// TIA Portal project "Pesteproject" (V15.1) (continued)
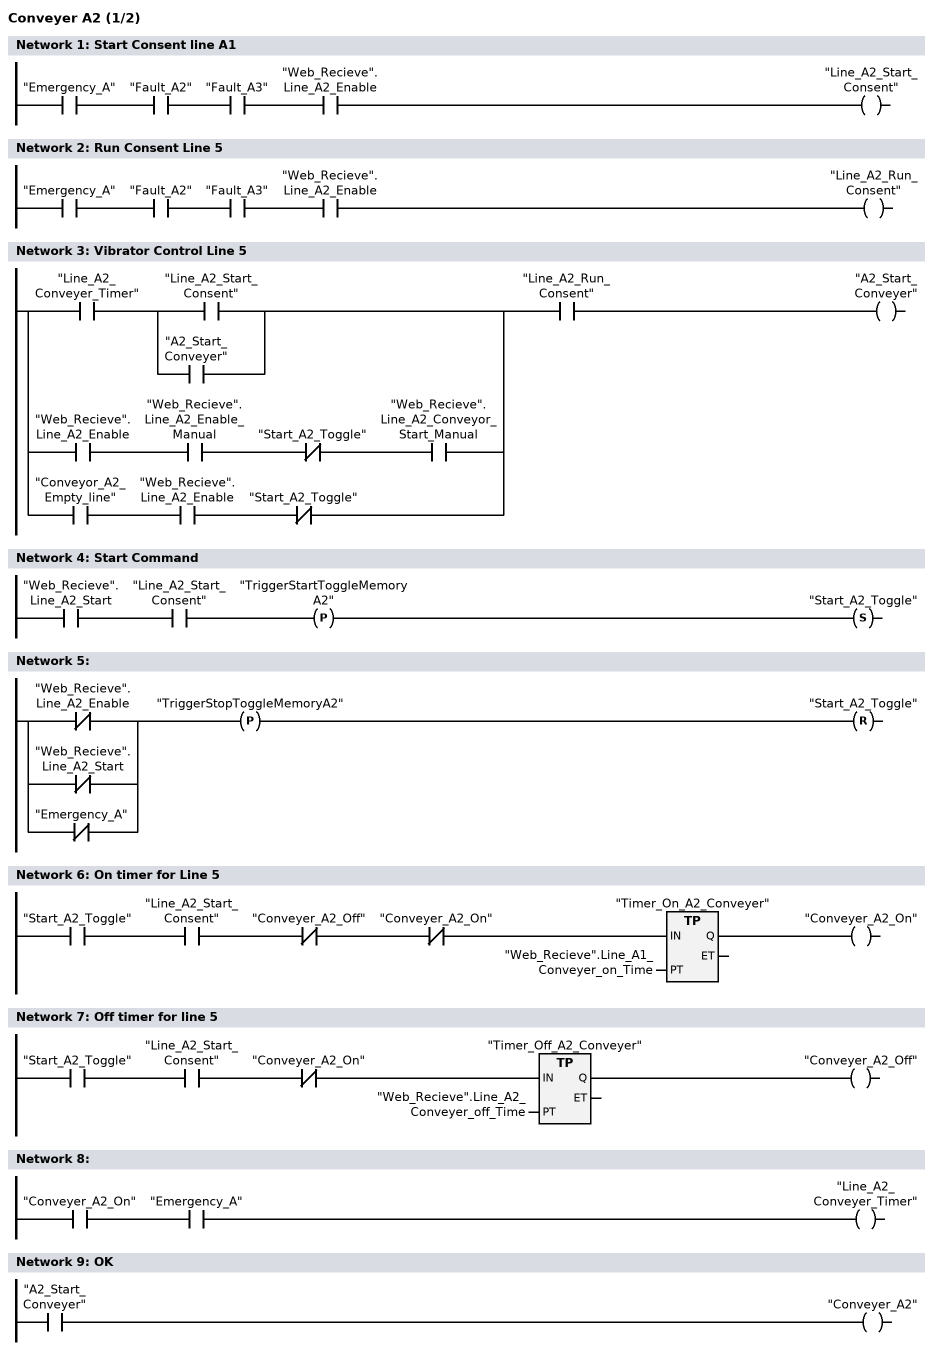
   RUNG wire#powerrail
      Contact( "Emergency_A" )
      Contact( "Fault_A2" )
      Contact( "Fault_A3" )
      Contact( "Web_Recieve".Line_A2_Enable )
      Coil( "Line_A2_Start_Consent" )
   END_RUNG
   // the same network as SCL:
   "Line_A2_Start_Consent" := "Emergency_A" AND "Fault_A2" AND "Fault_A3" AND "Web_Recieve".Line_A2_Enable;
END_REGION

REGION Network 2: Run Consent Line 5
   RUNG wire#powerrail
      Contact( "Emergency_A" )
      Contact( "Fault_A2" )
      Contact( "Fault_A3" )
      Contact( "Web_Recieve".Line_A2_Enable )
      Coil( "Line_A2_Run_Consent" )
   END_RUNG
   // the same network as SCL:
   "Line_A2_Run_Consent" := "Emergency_A" AND "Fault_A2" AND "Fault_A3" AND "Web_Recieve".Line_A2_Enable;
END_REGION

REGION Network 3: Vibrator Control Line 5
   RUNG wire#powerrail
      Contact( "Line_A2_Conveyer_Timer" )
      wire#w1
      Contact( "Line_A2_Start_Consent" )
      wire#w2
      Contact( "Line_A2_Run_Consent" )
      Coil( "A2_Start_Conveyer" )
   END_RUNG
   RUNG wire#w1
      Contact( "A2_Start_Conveyer" )
   END_RUNG wire#w2
   RUNG wire#powerrail
      Contact( "Web_Recieve".Line_A2_Enable )
      Contact( "Web_Recieve".Line_A2_Enable_Manual )
      I_Contact( "Start_A2_Toggle" )
      Contact( "Web_Recieve".Line_A2_Conveyor_Start_Manual )
   END_RUNG wire#w2
   RUNG wire#powerrail
      Contact( "Conveyor_A2_Empty_line" )
      Contact( "Web_Recieve".Line_A2_Enable )
      I_Contact( "Start_A2_Toggle" )
   END_RUNG wire#w2
   // the same network as SCL:
   "A2_Start_Conveyer" := (("Line_A2_Conveyer_Timer" AND ("Line_A2_Start_Consent" OR "A2_Start_Conveyer")) OR ("Web_Recieve".Line_A2_Enable AND "Web_Recieve".Line_A2_Enable_Manual AND NOT "Start_A2_Toggle" AND "Web_Recieve".Line_A2_Conveyor_Start_Manual) OR ("Conveyor_A2_Empty_line" AND "Web_Recieve".Line_A2_Enable AND NOT "Start_A2_Toggle")) AND "Line_A2_Run_Consent";
END_REGION

REGION Network 4: Start Command
   RUNG wire#powerrail
      Contact( "Web_Recieve".Line_A2_Start )
      Contact( "Line_A2_Start_Consent" )
      P_Trig( "TriggerStartToggleMemoryA2" )
      S_Coil( "Start_A2_Toggle" )
   END_RUNG
   // the same network as SCL:
   #_w1 := "Web_Recieve".Line_A2_Start AND "Line_A2_Start_Consent";
   #_w2 := #_w1 AND NOT "TriggerStartToggleMemoryA2";   // rising edge
   "TriggerStartToggleMemoryA2" := #_w1;
   IF #_w2 THEN "Start_A2_Toggle" := TRUE; END_IF;
END_REGION

REGION Network 5
   RUNG wire#powerrail
      I_Contact( "Web_Recieve".Line_A2_Enable )
      wire#w1
      P_Trig( "TriggerStopToggleMemoryA2" )
      R_Coil( "Start_A2_Toggle" )
   END_RUNG
   RUNG wire#powerrail
      I_Contact( "Web_Recieve".Line_A2_Start )
   END_RUNG wire#w1
   RUNG wire#powerrail
      I_Contact( "Emergency_A" )
   END_RUNG wire#w1
   // the same network as SCL:
   #_w1 := NOT "Web_Recieve".Line_A2_Enable OR NOT "Web_Recieve".Line_A2_Start OR NOT "Emergency_A";
   #_w2 := #_w1 AND NOT "TriggerStopToggleMemoryA2";   // rising edge
   "TriggerStopToggleMemoryA2" := #_w1;
   IF #_w2 THEN "Start_A2_Toggle" := FALSE; END_IF;
END_REGION

REGION Network 6: On timer for Line 5
   "Timer_On_A2_Conveyer".TP(IN := "Start_A2_Toggle" AND "Line_A2_Start_Consent" AND NOT "Conveyer_A2_Off" AND NOT "Conveyer_A2_On",
                           PT := "Web_Recieve".Line_A1_Conveyer_on_Time);
   "Conveyer_A2_On" := "Timer_On_A2_Conveyer".Q;
END_REGION

REGION Network 7: Off timer for line 5
   "Timer_Off_A2_Conveyer".TP(IN := "Start_A2_Toggle" AND "Line_A2_Start_Consent" AND NOT "Conveyer_A2_On",
                           PT := "Web_Recieve".Line_A2_Conveyer_off_Time);
   "Conveyer_A2_Off" := "Timer_Off_A2_Conveyer".Q;
END_REGION

REGION Network 8
   RUNG wire#powerrail
      Contact( "Conveyer_A2_On" )
      Contact( "Emergency_A" )
      Coil( "Line_A2_Conveyer_Timer" )
   END_RUNG
   // the same network as SCL:
   "Line_A2_Conveyer_Timer" := "Conveyer_A2_On" AND "Emergency_A";
END_REGION

REGION Network 9: OK
   RUNG wire#powerrail
      Contact( "A2_Start_Conveyer" )
      Coil( "Conveyer_A2" )
   END_RUNG
   // the same network as SCL:
   "Conveyer_A2" := "A2_Start_Conveyer";
END_REGION

REGION Network 10: emergency or stop or disable reser Timers
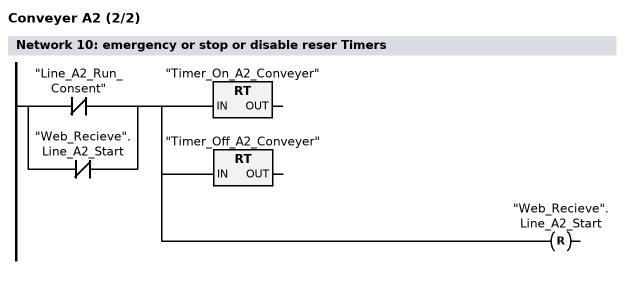
   RUNG wire#powerrail
      I_Contact( "Line_A2_Run_Consent" )
      wire#w1
      RT_Coil( "Timer_On_A2_Conveyer" )
   END_RUNG
   RUNG wire#powerrail
      I_Contact( "Web_Recieve".Line_A2_Start )
   END_RUNG wire#w1
   RUNG wire#w1
      RT_Coil( "Timer_Off_A2_Conveyer" )
   END_RUNG
   RUNG wire#w1
      R_Coil( "Web_Recieve".Line_A2_Start )
   END_RUNG
   // the same network as SCL:
   #_w1 := NOT "Line_A2_Run_Consent" OR NOT "Web_Recieve".Line_A2_Start;
   IF #_w1 THEN
       RESET_TIMER("Timer_On_A2_Conveyer");
       RESET_TIMER("Timer_Off_A2_Conveyer");
       "Web_Recieve".Line_A2_Start := FALSE;
   END_IF;
END_REGION
END_FUNCTION_BLOCK

FUNCTION_BLOCK "Conveyer B1"   // FB3, LAD
{ S7_Optimized_Access := 'TRUE' }
VERSION : 0.1
   VAR_TEMP   // added for the SCL form of the ladder/FBD networks
      _w1 : Bool;
      _w2 : Bool;
   END_VAR
BEGIN

REGION Network 1: Start Consent line A1
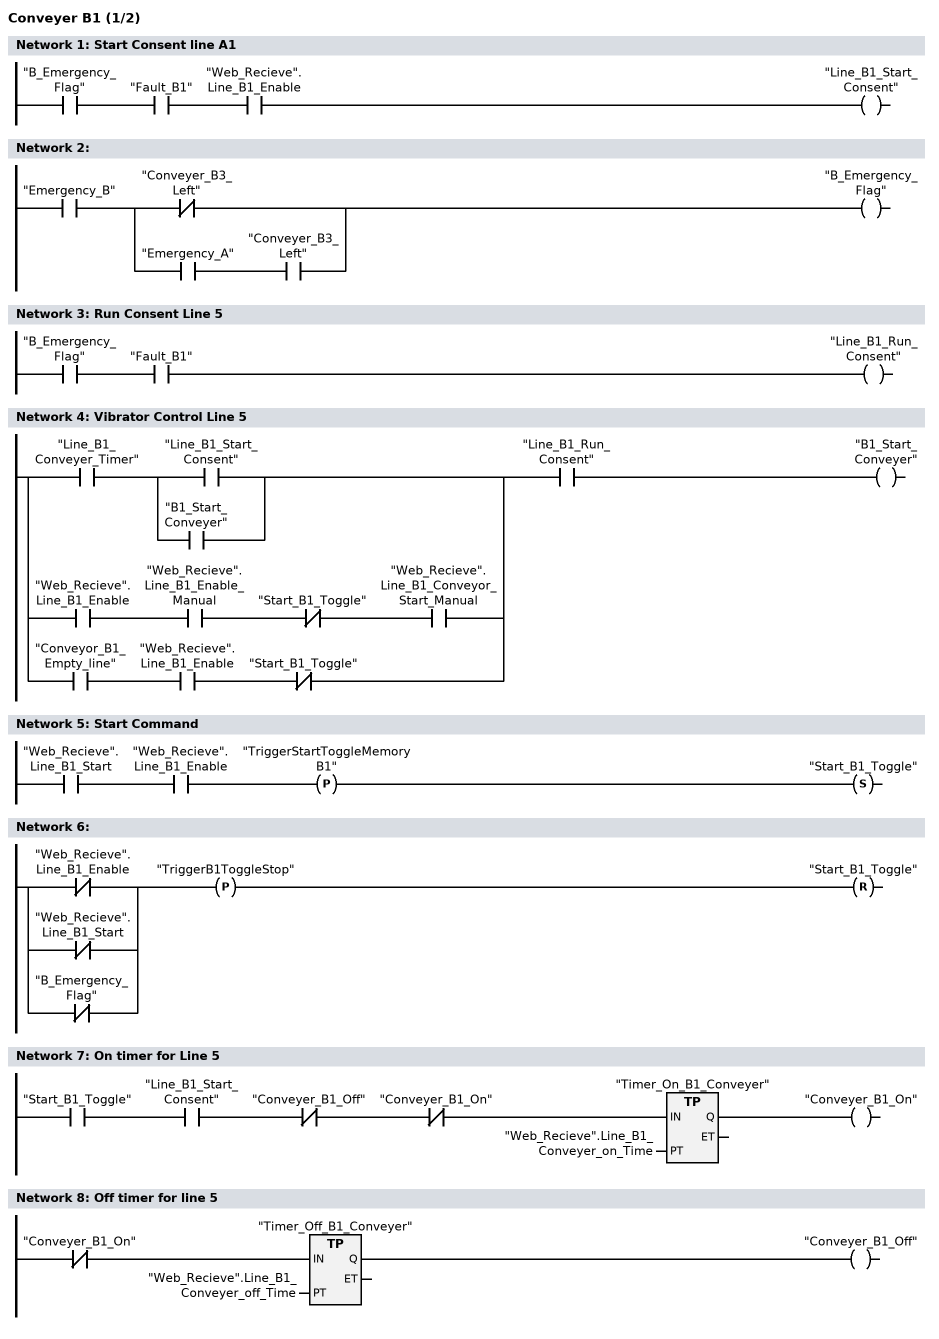
   RUNG wire#powerrail
      Contact( "B_Emergency_Flag" )
      Contact( "Fault_B1" )
      Contact( "Web_Recieve".Line_B1_Enable )
      Coil( "Line_B1_Start_Consent" )
   END_RUNG
   // the same network as SCL:
   "Line_B1_Start_Consent" := "B_Emergency_Flag" AND "Fault_B1" AND "Web_Recieve".Line_B1_Enable;
END_REGION

REGION Network 2
   RUNG wire#powerrail
      Contact( "Emergency_B" )
      wire#w1
      I_Contact( "Conveyer_B3_Left" )
      wire#w2
      Coil( "B_Emergency_Flag" )
   END_RUNG
   RUNG wire#w1
      Contact( "Emergency_A" )
      Contact( "Conveyer_B3_Left" )
   END_RUNG wire#w2
   // the same network as SCL:
   "B_Emergency_Flag" := "Emergency_B" AND (NOT "Conveyer_B3_Left" OR ("Emergency_A" AND "Conveyer_B3_Left"));
END_REGION

REGION Network 3: Run Consent Line 5
   RUNG wire#powerrail
      Contact( "B_Emergency_Flag" )
      Contact( "Fault_B1" )
      Coil( "Line_B1_Run_Consent" )
   END_RUNG
   // the same network as SCL:
   "Line_B1_Run_Consent" := "B_Emergency_Flag" AND "Fault_B1";
END_REGION

REGION Network 4: Vibrator Control Line 5
   RUNG wire#powerrail
      Contact( "Line_B1_Conveyer_Timer" )
      wire#w1
      Contact( "Line_B1_Start_Consent" )
      wire#w2
      Contact( "Line_B1_Run_Consent" )
      Coil( "B1_Start_Conveyer" )
   END_RUNG
   RUNG wire#w1
      Contact( "B1_Start_Conveyer" )
   END_RUNG wire#w2
   RUNG wire#powerrail
      Contact( "Web_Recieve".Line_B1_Enable )
      Contact( "Web_Recieve".Line_B1_Enable_Manual )
      I_Contact( "Start_B1_Toggle" )
      Contact( "Web_Recieve".Line_B1_Conveyor_Start_Manual )
   END_RUNG wire#w2
   RUNG wire#powerrail
      Contact( "Conveyor_B1_Empty_line" )
      Contact( "Web_Recieve".Line_B1_Enable )
      I_Contact( "Start_B1_Toggle" )
   END_RUNG wire#w2
   // the same network as SCL:
   "B1_Start_Conveyer" := (("Line_B1_Conveyer_Timer" AND ("Line_B1_Start_Consent" OR "B1_Start_Conveyer")) OR ("Web_Recieve".Line_B1_Enable AND "Web_Recieve".Line_B1_Enable_Manual AND NOT "Start_B1_Toggle" AND "Web_Recieve".Line_B1_Conveyor_Start_Manual) OR ("Conveyor_B1_Empty_line" AND "Web_Recieve".Line_B1_Enable AND NOT "Start_B1_Toggle")) AND "Line_B1_Run_Consent";
END_REGION

REGION Network 5: Start Command
   RUNG wire#powerrail
      Contact( "Web_Recieve".Line_B1_Start )
      Contact( "Web_Recieve".Line_B1_Enable )
      P_Trig( "TriggerStartToggleMemoryB1" )
      S_Coil( "Start_B1_Toggle" )
   END_RUNG
   // the same network as SCL:
   #_w1 := "Web_Recieve".Line_B1_Start AND "Web_Recieve".Line_B1_Enable;
   #_w2 := #_w1 AND NOT "TriggerStartToggleMemoryB1";   // rising edge
   "TriggerStartToggleMemoryB1" := #_w1;
   IF #_w2 THEN "Start_B1_Toggle" := TRUE; END_IF;
END_REGION

REGION Network 6
   RUNG wire#powerrail
      I_Contact( "Web_Recieve".Line_B1_Enable )
      wire#w1
      P_Trig( "TriggerB1ToggleStop" )
      R_Coil( "Start_B1_Toggle" )
   END_RUNG
   RUNG wire#powerrail
      I_Contact( "Web_Recieve".Line_B1_Start )
   END_RUNG wire#w1
   RUNG wire#powerrail
      I_Contact( "B_Emergency_Flag" )
   END_RUNG wire#w1
   // the same network as SCL:
   #_w1 := NOT "Web_Recieve".Line_B1_Enable OR NOT "Web_Recieve".Line_B1_Start OR NOT "B_Emergency_Flag";
   #_w2 := #_w1 AND NOT "TriggerB1ToggleStop";   // rising edge
   "TriggerB1ToggleStop" := #_w1;
   IF #_w2 THEN "Start_B1_Toggle" := FALSE; END_IF;
END_REGION

REGION Network 7: On timer for Line 5
   "Timer_On_B1_Conveyer".TP(IN := "Start_B1_Toggle" AND "Line_B1_Start_Consent" AND NOT "Conveyer_B1_Off" AND NOT "Conveyer_B1_On",
                           PT := "Web_Recieve".Line_B1_Conveyer_on_Time);
   "Conveyer_B1_On" := "Timer_On_B1_Conveyer".Q;
END_REGION

REGION Network 8: Off timer for line 5
   "Timer_Off_B1_Conveyer".TP(IN := NOT "Conveyer_B1_On", PT := "Web_Recieve".Line_B1_Conveyer_off_Time);
   "Conveyer_B1_Off" := "Timer_Off_B1_Conveyer".Q;
END_REGION

REGION Network 9
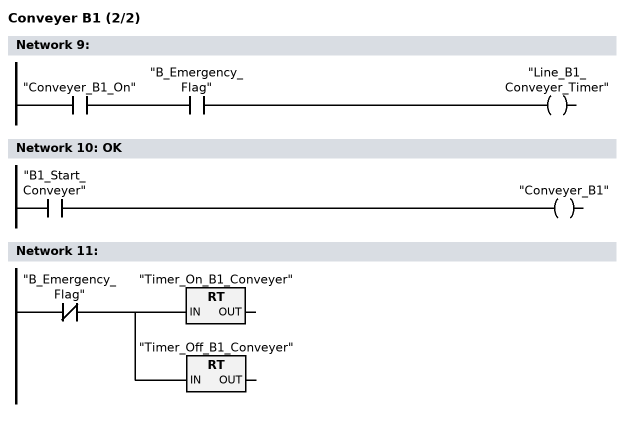
   RUNG wire#powerrail
      Contact( "Conveyer_B1_On" )
      Contact( "B_Emergency_Flag" )
      Coil( "Line_B1_Conveyer_Timer" )
   END_RUNG
   // the same network as SCL:
   "Line_B1_Conveyer_Timer" := "Conveyer_B1_On" AND "B_Emergency_Flag";
END_REGION

REGION Network 10: OK
   RUNG wire#powerrail
      Contact( "B1_Start_Conveyer" )
      Coil( "Conveyer_B1" )
   END_RUNG
   // the same network as SCL:
   "Conveyer_B1" := "B1_Start_Conveyer";
END_REGION

REGION Network 11
   RUNG wire#powerrail
      I_Contact( "B_Emergency_Flag" )
      wire#w1
      RT_Coil( "Timer_On_B1_Conveyer" )
   END_RUNG
   RUNG wire#w1
      RT_Coil( "Timer_Off_B1_Conveyer" )
   END_RUNG
   // the same network as SCL:
   IF NOT "B_Emergency_Flag" THEN
       RESET_TIMER("Timer_On_B1_Conveyer");
       RESET_TIMER("Timer_Off_B1_Conveyer");
   END_IF;
END_REGION
END_FUNCTION_BLOCK

FUNCTION_BLOCK "Conveyer B2"   // FB4, LAD
{ S7_Optimized_Access := 'TRUE' }
VERSION : 0.1
   VAR_TEMP   // added for the SCL form of the ladder/FBD networks
      _w1 : Bool;
      _w2 : Bool;
   END_VAR
BEGIN

REGION Network 1: Start Consent line A1
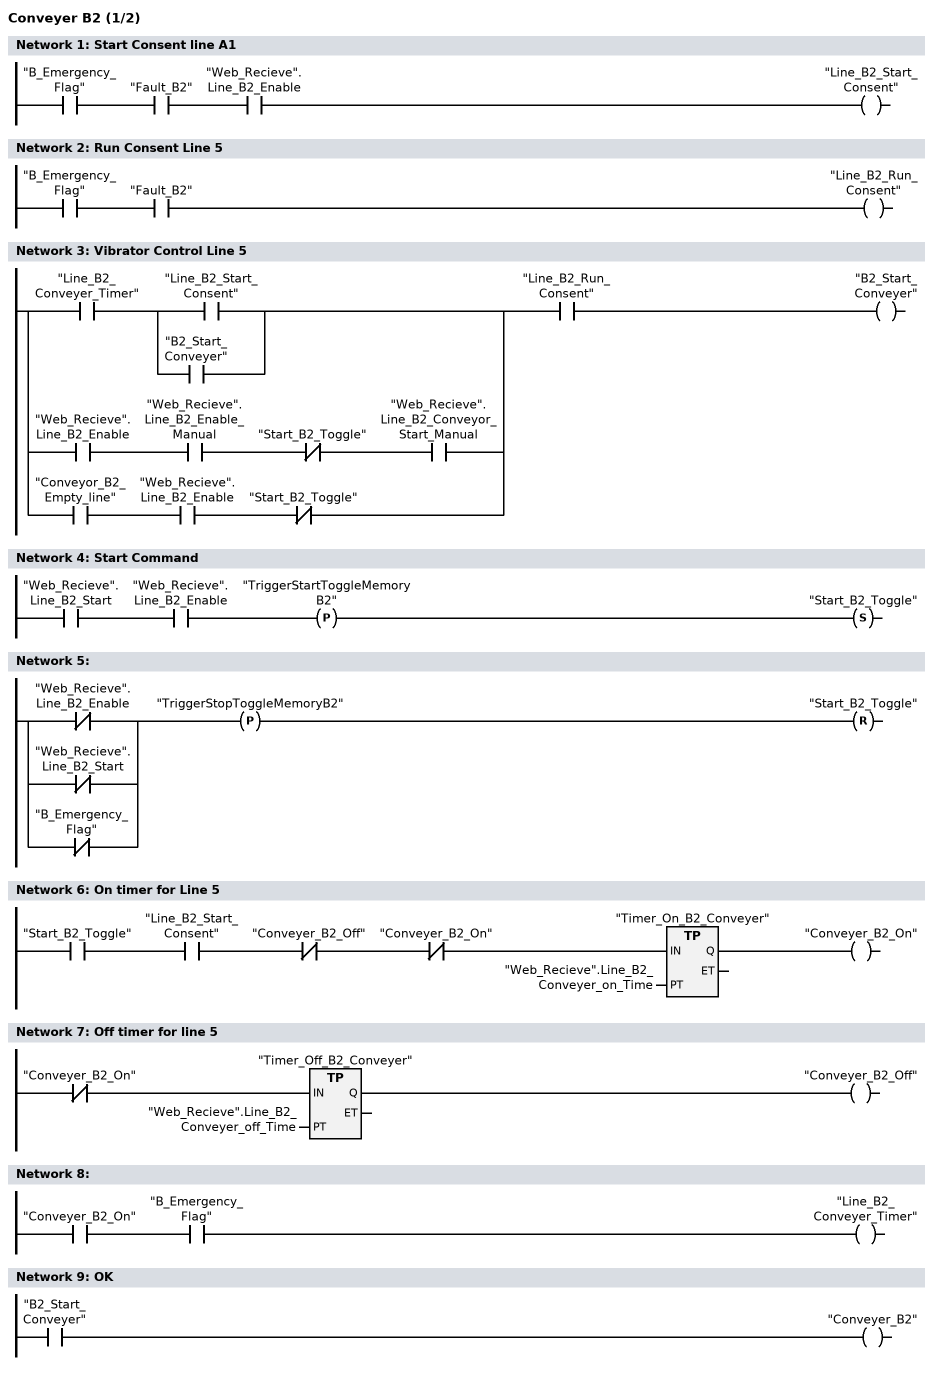
   RUNG wire#powerrail
      Contact( "B_Emergency_Flag" )
      Contact( "Fault_B2" )
      Contact( "Web_Recieve".Line_B2_Enable )
      Coil( "Line_B2_Start_Consent" )
   END_RUNG
   // the same network as SCL:
   "Line_B2_Start_Consent" := "B_Emergency_Flag" AND "Fault_B2" AND "Web_Recieve".Line_B2_Enable;
END_REGION

REGION Network 2: Run Consent Line 5
   RUNG wire#powerrail
      Contact( "B_Emergency_Flag" )
      Contact( "Fault_B2" )
      Coil( "Line_B2_Run_Consent" )
   END_RUNG
   // the same network as SCL:
   "Line_B2_Run_Consent" := "B_Emergency_Flag" AND "Fault_B2";
END_REGION

REGION Network 3: Vibrator Control Line 5
   RUNG wire#powerrail
      Contact( "Line_B2_Conveyer_Timer" )
      wire#w1
      Contact( "Line_B2_Start_Consent" )
      wire#w2
      Contact( "Line_B2_Run_Consent" )
      Coil( "B2_Start_Conveyer" )
   END_RUNG
   RUNG wire#w1
      Contact( "B2_Start_Conveyer" )
   END_RUNG wire#w2
   RUNG wire#powerrail
      Contact( "Web_Recieve".Line_B2_Enable )
      Contact( "Web_Recieve".Line_B2_Enable_Manual )
      I_Contact( "Start_B2_Toggle" )
      Contact( "Web_Recieve".Line_B2_Conveyor_Start_Manual )
   END_RUNG wire#w2
   RUNG wire#powerrail
      Contact( "Conveyor_B2_Empty_line" )
      Contact( "Web_Recieve".Line_B2_Enable )
      I_Contact( "Start_B2_Toggle" )
   END_RUNG wire#w2
   // the same network as SCL:
   "B2_Start_Conveyer" := (("Line_B2_Conveyer_Timer" AND ("Line_B2_Start_Consent" OR "B2_Start_Conveyer")) OR ("Web_Recieve".Line_B2_Enable AND "Web_Recieve".Line_B2_Enable_Manual AND NOT "Start_B2_Toggle" AND "Web_Recieve".Line_B2_Conveyor_Start_Manual) OR ("Conveyor_B2_Empty_line" AND "Web_Recieve".Line_B2_Enable AND NOT "Start_B2_Toggle")) AND "Line_B2_Run_Consent";
END_REGION

REGION Network 4: Start Command
   RUNG wire#powerrail
      Contact( "Web_Recieve".Line_B2_Start )
      Contact( "Web_Recieve".Line_B2_Enable )
      P_Trig( "TriggerStartToggleMemoryB2" )
      S_Coil( "Start_B2_Toggle" )
   END_RUNG
   // the same network as SCL:
   #_w1 := "Web_Recieve".Line_B2_Start AND "Web_Recieve".Line_B2_Enable;
   #_w2 := #_w1 AND NOT "TriggerStartToggleMemoryB2";   // rising edge
   "TriggerStartToggleMemoryB2" := #_w1;
   IF #_w2 THEN "Start_B2_Toggle" := TRUE; END_IF;
END_REGION

REGION Network 5
   RUNG wire#powerrail
      I_Contact( "Web_Recieve".Line_B2_Enable )
      wire#w1
      P_Trig( "TriggerStopToggleMemoryB2" )
      R_Coil( "Start_B2_Toggle" )
   END_RUNG
   RUNG wire#powerrail
      I_Contact( "Web_Recieve".Line_B2_Start )
   END_RUNG wire#w1
   RUNG wire#powerrail
      I_Contact( "B_Emergency_Flag" )
   END_RUNG wire#w1
   // the same network as SCL:
   #_w1 := NOT "Web_Recieve".Line_B2_Enable OR NOT "Web_Recieve".Line_B2_Start OR NOT "B_Emergency_Flag";
   #_w2 := #_w1 AND NOT "TriggerStopToggleMemoryB2";   // rising edge
   "TriggerStopToggleMemoryB2" := #_w1;
   IF #_w2 THEN "Start_B2_Toggle" := FALSE; END_IF;
END_REGION

REGION Network 6: On timer for Line 5
   "Timer_On_B2_Conveyer".TP(IN := "Start_B2_Toggle" AND "Line_B2_Start_Consent" AND NOT "Conveyer_B2_Off" AND NOT "Conveyer_B2_On",
                           PT := "Web_Recieve".Line_B2_Conveyer_on_Time);
   "Conveyer_B2_On" := "Timer_On_B2_Conveyer".Q;
END_REGION

REGION Network 7: Off timer for line 5
   "Timer_Off_B2_Conveyer".TP(IN := NOT "Conveyer_B2_On", PT := "Web_Recieve".Line_B2_Conveyer_off_Time);
   "Conveyer_B2_Off" := "Timer_Off_B2_Conveyer".Q;
END_REGION

REGION Network 8
   RUNG wire#powerrail
      Contact( "Conveyer_B2_On" )
      Contact( "B_Emergency_Flag" )
      Coil( "Line_B2_Conveyer_Timer" )
   END_RUNG
   // the same network as SCL:
   "Line_B2_Conveyer_Timer" := "Conveyer_B2_On" AND "B_Emergency_Flag";
END_REGION

REGION Network 9: OK
   RUNG wire#powerrail
      Contact( "B2_Start_Conveyer" )
      Coil( "Conveyer_B2" )
   END_RUNG
   // the same network as SCL:
   "Conveyer_B2" := "B2_Start_Conveyer";
END_REGION

REGION Network 10
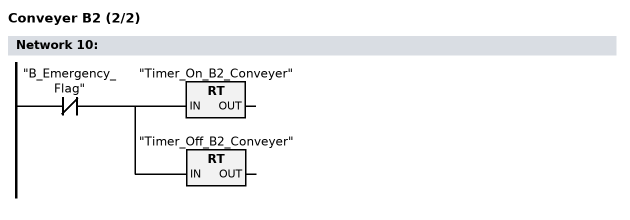
   RUNG wire#powerrail
      I_Contact( "B_Emergency_Flag" )
      wire#w1
      RT_Coil( "Timer_On_B2_Conveyer" )
   END_RUNG
   RUNG wire#w1
      RT_Coil( "Timer_Off_B2_Conveyer" )
   END_RUNG
   // the same network as SCL:
   IF NOT "B_Emergency_Flag" THEN
       RESET_TIMER("Timer_On_B2_Conveyer");
       RESET_TIMER("Timer_Off_B2_Conveyer");
   END_IF;
END_REGION
END_FUNCTION_BLOCK

FUNCTION_BLOCK "Vibrator A1"   // FB5, LAD
{ S7_Optimized_Access := 'TRUE' }
VERSION : 0.1
   VAR_TEMP
      RemainTime : DInt;
   END_VAR
BEGIN

REGION Network 1
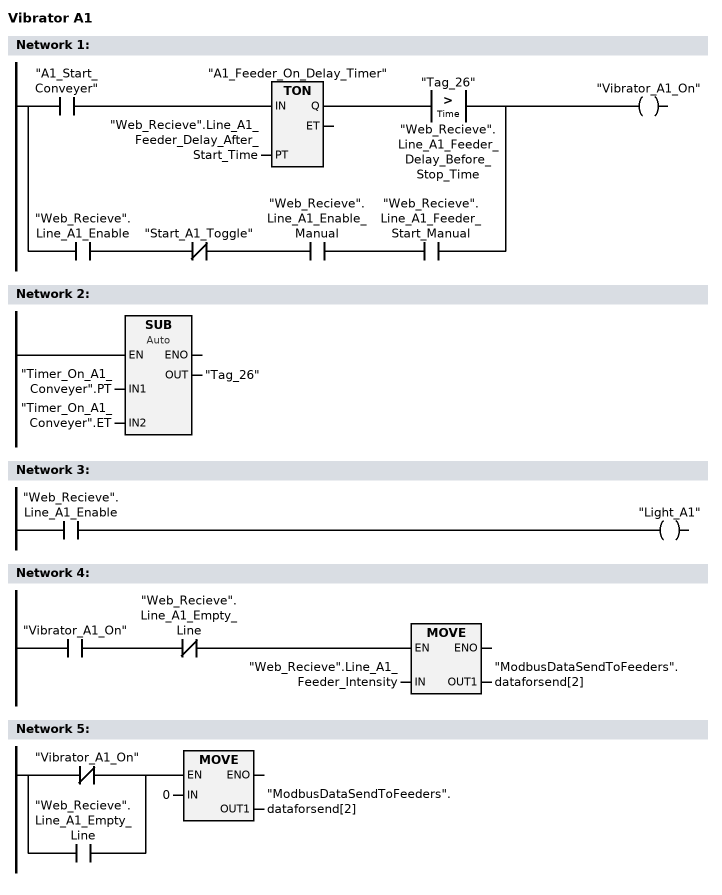
   "A1_Feeder_On_Delay_Timer".TON(IN := "A1_Start_Conveyer",
                           PT := "Web_Recieve".Line_A1_Feeder_Delay_After_Start_Time);
   "Vibrator_A1_On" := ("A1_Feeder_On_Delay_Timer".Q AND ("Tag_26" > "Web_Recieve".Line_A1_Feeder_Delay_Before_Stop_Time)) OR ("Web_Recieve".Line_A1_Enable AND NOT "Start_A1_Toggle" AND "Web_Recieve".Line_A1_Enable_Manual AND "Web_Recieve".Line_A1_Feeder_Start_Manual);
END_REGION

REGION Network 2
   RUNG wire#powerrail
      Sub(in1 := "Timer_On_A1_Conveyer".PT, in2 := "Timer_On_A1_Conveyer".ET, out => "Tag_26")
   END_RUNG
   // the same network as SCL:
   "Tag_26" := "Timer_On_A1_Conveyer".PT - "Timer_On_A1_Conveyer".ET;
END_REGION

REGION Network 3
   RUNG wire#powerrail
      Contact( "Web_Recieve".Line_A1_Enable )
      Coil( "Light_A1" )
   END_RUNG
   // the same network as SCL:
   "Light_A1" := "Web_Recieve".Line_A1_Enable;
END_REGION

REGION Network 4
   RUNG wire#powerrail
      Contact( "Vibrator_A1_On" )
      I_Contact( "Web_Recieve".Line_A1_Empty_Line )
      Move(in := "Web_Recieve".Line_A1_Feeder_Intensity, out1 => "ModbusDataSendToFeeders".dataforsend[2])
   END_RUNG
   // the same network as SCL:
   IF "Vibrator_A1_On" AND NOT "Web_Recieve".Line_A1_Empty_Line THEN
       "ModbusDataSendToFeeders".dataforsend[2] := "Web_Recieve".Line_A1_Feeder_Intensity;
   END_IF;
END_REGION

REGION Network 5
   RUNG wire#powerrail
      I_Contact( "Vibrator_A1_On" )
      wire#w1
      Move(in := 0, out1 => "ModbusDataSendToFeeders".dataforsend[2])
   END_RUNG
   RUNG wire#powerrail
      Contact( "Web_Recieve".Line_A1_Empty_Line )
   END_RUNG wire#w1
   // the same network as SCL:
   IF NOT "Vibrator_A1_On" OR "Web_Recieve".Line_A1_Empty_Line THEN
       "ModbusDataSendToFeeders".dataforsend[2] := 0;
   END_IF;
END_REGION
END_FUNCTION_BLOCK

FUNCTION_BLOCK "Vibrator A2"   // FB6, LAD
{ S7_Optimized_Access := 'TRUE' }
VERSION : 0.1
BEGIN

REGION Network 1
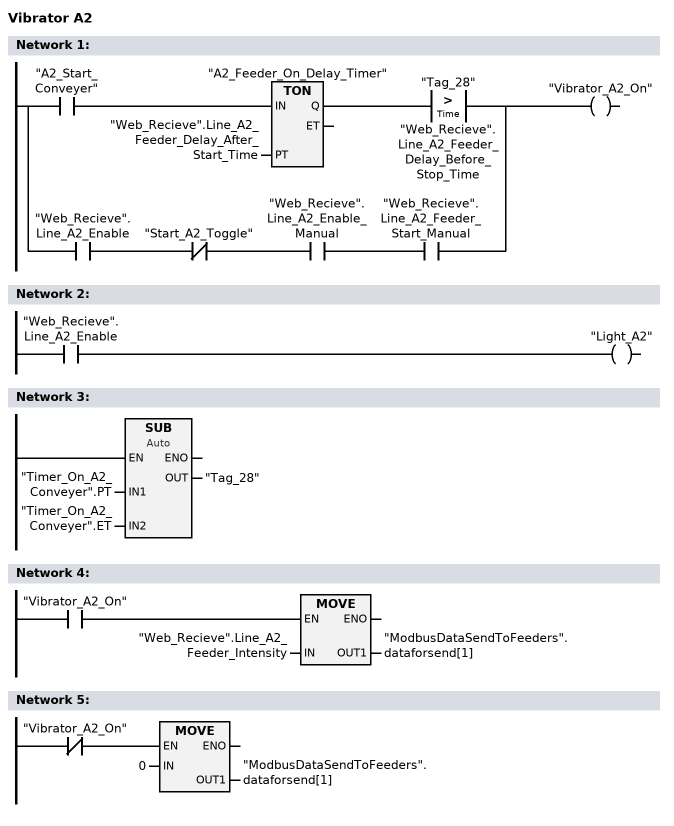
   "A2_Feeder_On_Delay_Timer".TON(IN := "A2_Start_Conveyer",
                           PT := "Web_Recieve".Line_A2_Feeder_Delay_After_Start_Time);
   "Vibrator_A2_On" := ("A2_Feeder_On_Delay_Timer".Q AND ("Tag_28" > "Web_Recieve".Line_A2_Feeder_Delay_Before_Stop_Time)) OR ("Web_Recieve".Line_A2_Enable AND NOT "Start_A2_Toggle" AND "Web_Recieve".Line_A2_Enable_Manual AND "Web_Recieve".Line_A2_Feeder_Start_Manual);
END_REGION

REGION Network 2
   RUNG wire#powerrail
      Contact( "Web_Recieve".Line_A2_Enable )
      Coil( "Light_A2" )
   END_RUNG
   // the same network as SCL:
   "Light_A2" := "Web_Recieve".Line_A2_Enable;
END_REGION

REGION Network 3
   RUNG wire#powerrail
      Sub(in1 := "Timer_On_A2_Conveyer".PT, in2 := "Timer_On_A2_Conveyer".ET, out => "Tag_28")
   END_RUNG
   // the same network as SCL:
   "Tag_28" := "Timer_On_A2_Conveyer".PT - "Timer_On_A2_Conveyer".ET;
END_REGION

REGION Network 4
   RUNG wire#powerrail
      Contact( "Vibrator_A2_On" )
      Move(in := "Web_Recieve".Line_A2_Feeder_Intensity, out1 => "ModbusDataSendToFeeders".dataforsend[1])
   END_RUNG
   // the same network as SCL:
   IF "Vibrator_A2_On" THEN
       "ModbusDataSendToFeeders".dataforsend[1] := "Web_Recieve".Line_A2_Feeder_Intensity;
   END_IF;
END_REGION

REGION Network 5
   RUNG wire#powerrail
      I_Contact( "Vibrator_A2_On" )
      Move(in := 0, out1 => "ModbusDataSendToFeeders".dataforsend[1])
   END_RUNG
   // the same network as SCL:
   IF NOT "Vibrator_A2_On" THEN "ModbusDataSendToFeeders".dataforsend[1] := 0; END_IF;
END_REGION
END_FUNCTION_BLOCK

FUNCTION_BLOCK "Vibrator B1"   // FB7, LAD
{ S7_Optimized_Access := 'TRUE' }
VERSION : 0.1
BEGIN

REGION Network 1
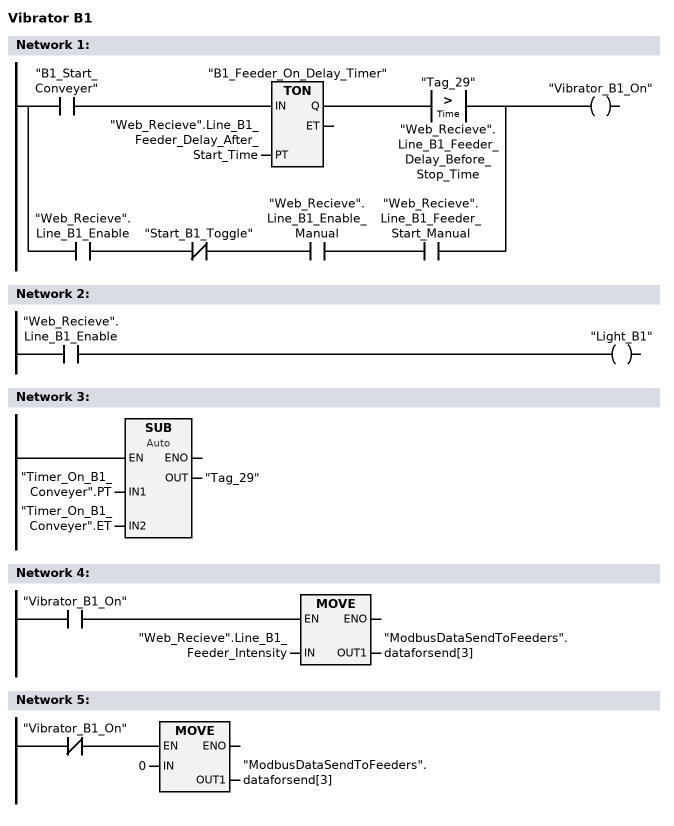
   "B1_Feeder_On_Delay_Timer".TON(IN := "B1_Start_Conveyer",
                           PT := "Web_Recieve".Line_B1_Feeder_Delay_After_Start_Time);
   "Vibrator_B1_On" := ("B1_Feeder_On_Delay_Timer".Q AND ("Tag_29" > "Web_Recieve".Line_B1_Feeder_Delay_Before_Stop_Time)) OR ("Web_Recieve".Line_B1_Enable AND NOT "Start_B1_Toggle" AND "Web_Recieve".Line_B1_Enable_Manual AND "Web_Recieve".Line_B1_Feeder_Start_Manual);
END_REGION

REGION Network 2
   RUNG wire#powerrail
      Contact( "Web_Recieve".Line_B1_Enable )
      Coil( "Light_B1" )
   END_RUNG
   // the same network as SCL:
   "Light_B1" := "Web_Recieve".Line_B1_Enable;
END_REGION

REGION Network 3
   RUNG wire#powerrail
      Sub(in1 := "Timer_On_B1_Conveyer".PT, in2 := "Timer_On_B1_Conveyer".ET, out => "Tag_29")
   END_RUNG
   // the same network as SCL:
   "Tag_29" := "Timer_On_B1_Conveyer".PT - "Timer_On_B1_Conveyer".ET;
END_REGION

REGION Network 4
   RUNG wire#powerrail
      Contact( "Vibrator_B1_On" )
      Move(in := "Web_Recieve".Line_B1_Feeder_Intensity, out1 => "ModbusDataSendToFeeders".dataforsend[3])
   END_RUNG
   // the same network as SCL:
   IF "Vibrator_B1_On" THEN
       "ModbusDataSendToFeeders".dataforsend[3] := "Web_Recieve".Line_B1_Feeder_Intensity;
   END_IF;
END_REGION

REGION Network 5
   RUNG wire#powerrail
      I_Contact( "Vibrator_B1_On" )
      Move(in := 0, out1 => "ModbusDataSendToFeeders".dataforsend[3])
   END_RUNG
   // the same network as SCL:
   IF NOT "Vibrator_B1_On" THEN "ModbusDataSendToFeeders".dataforsend[3] := 0; END_IF;
END_REGION
END_FUNCTION_BLOCK

FUNCTION_BLOCK "Vibrator B2"   // FB8, LAD
{ S7_Optimized_Access := 'TRUE' }
VERSION : 0.1
BEGIN

REGION Network 1
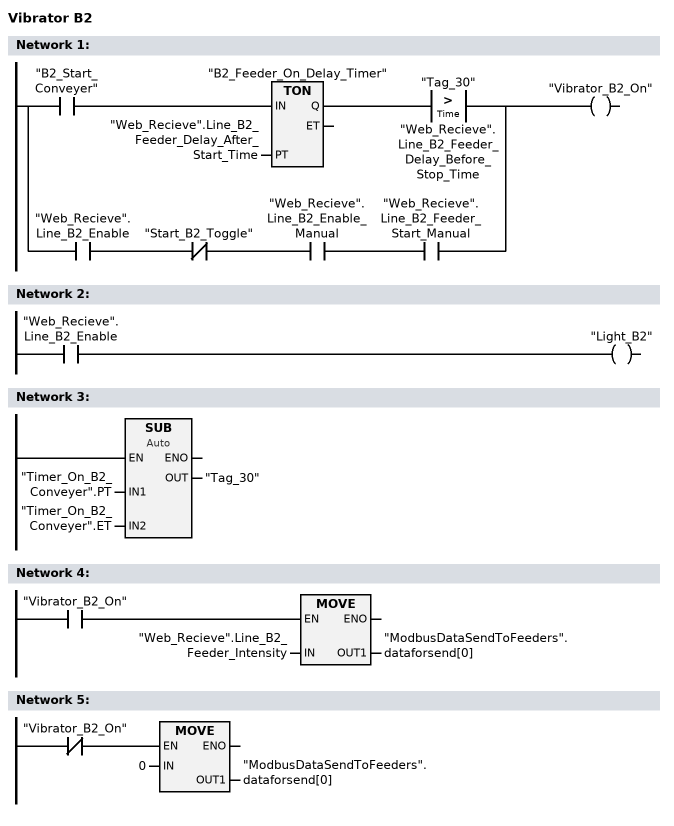
   "B2_Feeder_On_Delay_Timer".TON(IN := "B2_Start_Conveyer",
                           PT := "Web_Recieve".Line_B2_Feeder_Delay_After_Start_Time);
   "Vibrator_B2_On" := ("B2_Feeder_On_Delay_Timer".Q AND ("Tag_30" > "Web_Recieve".Line_B2_Feeder_Delay_Before_Stop_Time)) OR ("Web_Recieve".Line_B2_Enable AND NOT "Start_B2_Toggle" AND "Web_Recieve".Line_B2_Enable_Manual AND "Web_Recieve".Line_B2_Feeder_Start_Manual);
END_REGION

REGION Network 2
   RUNG wire#powerrail
      Contact( "Web_Recieve".Line_B2_Enable )
      Coil( "Light_B2" )
   END_RUNG
   // the same network as SCL:
   "Light_B2" := "Web_Recieve".Line_B2_Enable;
END_REGION

REGION Network 3
   RUNG wire#powerrail
      Sub(in1 := "Timer_On_B2_Conveyer".PT, in2 := "Timer_On_B2_Conveyer".ET, out => "Tag_30")
   END_RUNG
   // the same network as SCL:
   "Tag_30" := "Timer_On_B2_Conveyer".PT - "Timer_On_B2_Conveyer".ET;
END_REGION

REGION Network 4
   RUNG wire#powerrail
      Contact( "Vibrator_B2_On" )
      Move(in := "Web_Recieve".Line_B2_Feeder_Intensity, out1 => "ModbusDataSendToFeeders".dataforsend[0])
   END_RUNG
   // the same network as SCL:
   IF "Vibrator_B2_On" THEN
       "ModbusDataSendToFeeders".dataforsend[0] := "Web_Recieve".Line_B2_Feeder_Intensity;
   END_IF;
END_REGION

REGION Network 5
   RUNG wire#powerrail
      I_Contact( "Vibrator_B2_On" )
      Move(in := 0, out1 => "ModbusDataSendToFeeders".dataforsend[0])
   END_RUNG
   // the same network as SCL:
   IF NOT "Vibrator_B2_On" THEN "ModbusDataSendToFeeders".dataforsend[0] := 0; END_IF;
END_REGION
END_FUNCTION_BLOCK

FUNCTION_BLOCK "ConveyerA3_B3"   // FB9, LAD
{ S7_Optimized_Access := 'TRUE' }
VERSION : 0.1
BEGIN

REGION Network 1
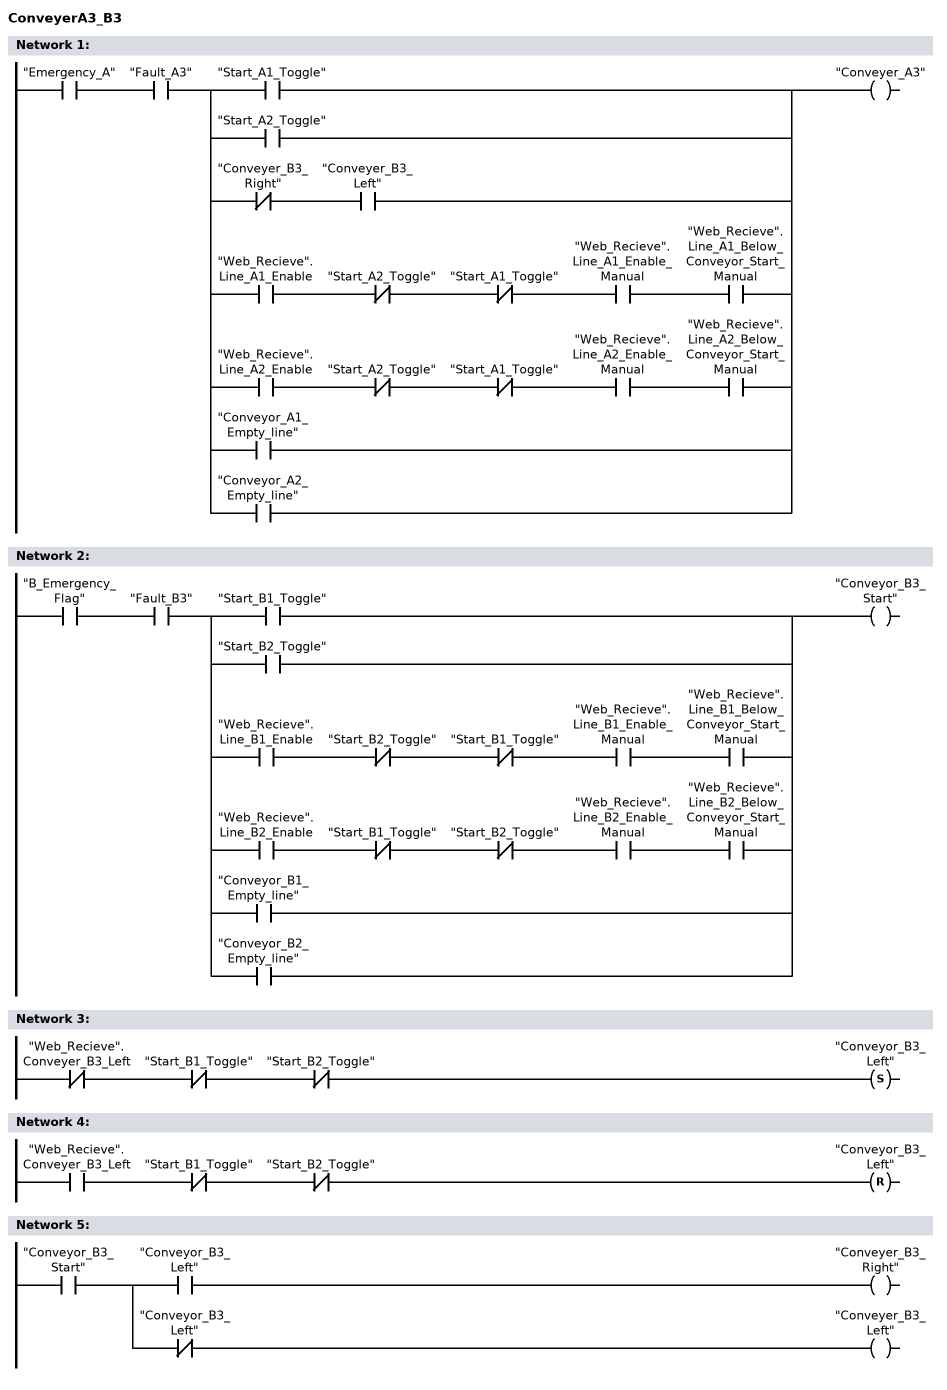
   RUNG wire#powerrail
      Contact( "Emergency_A" )
      Contact( "Fault_A3" )
      wire#w1
      Contact( "Start_A1_Toggle" )
      wire#w2
      Coil( "Conveyer_A3" )
   END_RUNG
   RUNG wire#w1
      Contact( "Start_A2_Toggle" )
   END_RUNG wire#w2
   RUNG wire#w1
      I_Contact( "Conveyer_B3_Right" )
      Contact( "Conveyer_B3_Left" )
   END_RUNG wire#w2
   RUNG wire#w1
      Contact( "Web_Recieve".Line_A1_Enable )
      I_Contact( "Start_A2_Toggle" )
      I_Contact( "Start_A1_Toggle" )
      Contact( "Web_Recieve".Line_A1_Enable_Manual )
      Contact( "Web_Recieve".Line_A1_Below_Conveyor_Start_Manual )
   END_RUNG wire#w2
   RUNG wire#w1
      Contact( "Web_Recieve".Line_A2_Enable )
      I_Contact( "Start_A2_Toggle" )
      I_Contact( "Start_A1_Toggle" )
      Contact( "Web_Recieve".Line_A2_Enable_Manual )
      Contact( "Web_Recieve".Line_A2_Below_Conveyor_Start_Manual )
   END_RUNG wire#w2
   RUNG wire#w1
      Contact( "Conveyor_A1_Empty_line" )
   END_RUNG wire#w2
   RUNG wire#w1
      Contact( "Conveyor_A2_Empty_line" )
   END_RUNG wire#w2
   // the same network as SCL:
   "Conveyer_A3" := "Emergency_A" AND "Fault_A3" AND ("Start_A1_Toggle" OR "Start_A2_Toggle" OR (NOT "Conveyer_B3_Right" AND "Conveyer_B3_Left") OR ("Web_Recieve".Line_A1_Enable AND NOT "Start_A2_Toggle" AND NOT "Start_A1_Toggle" AND "Web_Recieve".Line_A1_Enable_Manual AND "Web_Recieve".Line_A1_Below_Conveyor_Start_Manual) OR ("Web_Recieve".Line_A2_Enable AND NOT "Start_A2_Toggle" AND NOT "Start_A1_Toggle" AND "Web_Recieve".Line_A2_Enable_Manual AND "Web_Recieve".Line_A2_Below_Conveyor_Start_Manual) OR "Conveyor_A1_Empty_line" OR "Conveyor_A2_Empty_line");
END_REGION

REGION Network 2
   RUNG wire#powerrail
      Contact( "B_Emergency_Flag" )
      Contact( "Fault_B3" )
      wire#w1
      Contact( "Start_B1_Toggle" )
      wire#w2
      Coil( "Conveyor_B3_Start" )
   END_RUNG
   RUNG wire#w1
      Contact( "Start_B2_Toggle" )
   END_RUNG wire#w2
   RUNG wire#w1
      Contact( "Web_Recieve".Line_B1_Enable )
      I_Contact( "Start_B2_Toggle" )
      I_Contact( "Start_B1_Toggle" )
      Contact( "Web_Recieve".Line_B1_Enable_Manual )
      Contact( "Web_Recieve".Line_B1_Below_Conveyor_Start_Manual )
   END_RUNG wire#w2
   RUNG wire#w1
      Contact( "Web_Recieve".Line_B2_Enable )
      I_Contact( "Start_B1_Toggle" )
      I_Contact( "Start_B2_Toggle" )
      Contact( "Web_Recieve".Line_B2_Enable_Manual )
      Contact( "Web_Recieve".Line_B2_Below_Conveyor_Start_Manual )
   END_RUNG wire#w2
   RUNG wire#w1
      Contact( "Conveyor_B1_Empty_line" )
   END_RUNG wire#w2
   RUNG wire#w1
      Contact( "Conveyor_B2_Empty_line" )
   END_RUNG wire#w2
   // the same network as SCL:
   "Conveyor_B3_Start" := "B_Emergency_Flag" AND "Fault_B3" AND ("Start_B1_Toggle" OR "Start_B2_Toggle" OR ("Web_Recieve".Line_B1_Enable AND NOT "Start_B2_Toggle" AND NOT "Start_B1_Toggle" AND "Web_Recieve".Line_B1_Enable_Manual AND "Web_Recieve".Line_B1_Below_Conveyor_Start_Manual) OR ("Web_Recieve".Line_B2_Enable AND NOT "Start_B1_Toggle" AND NOT "Start_B2_Toggle" AND "Web_Recieve".Line_B2_Enable_Manual AND "Web_Recieve".Line_B2_Below_Conveyor_Start_Manual) OR "Conveyor_B1_Empty_line" OR "Conveyor_B2_Empty_line");
END_REGION

REGION Network 3
   RUNG wire#powerrail
      I_Contact( "Web_Recieve".Conveyer_B3_Left )
      I_Contact( "Start_B1_Toggle" )
      I_Contact( "Start_B2_Toggle" )
      S_Coil( "Conveyor_B3_Left" )
   END_RUNG
   // the same network as SCL:
   IF NOT "Web_Recieve".Conveyer_B3_Left AND NOT "Start_B1_Toggle" AND NOT "Start_B2_Toggle" THEN
       "Conveyor_B3_Left" := TRUE;
   END_IF;
END_REGION

REGION Network 4
   RUNG wire#powerrail
      Contact( "Web_Recieve".Conveyer_B3_Left )
      I_Contact( "Start_B1_Toggle" )
      I_Contact( "Start_B2_Toggle" )
      R_Coil( "Conveyor_B3_Left" )
   END_RUNG
   // the same network as SCL:
   IF "Web_Recieve".Conveyer_B3_Left AND NOT "Start_B1_Toggle" AND NOT "Start_B2_Toggle" THEN
       "Conveyor_B3_Left" := FALSE;
   END_IF;
END_REGION
